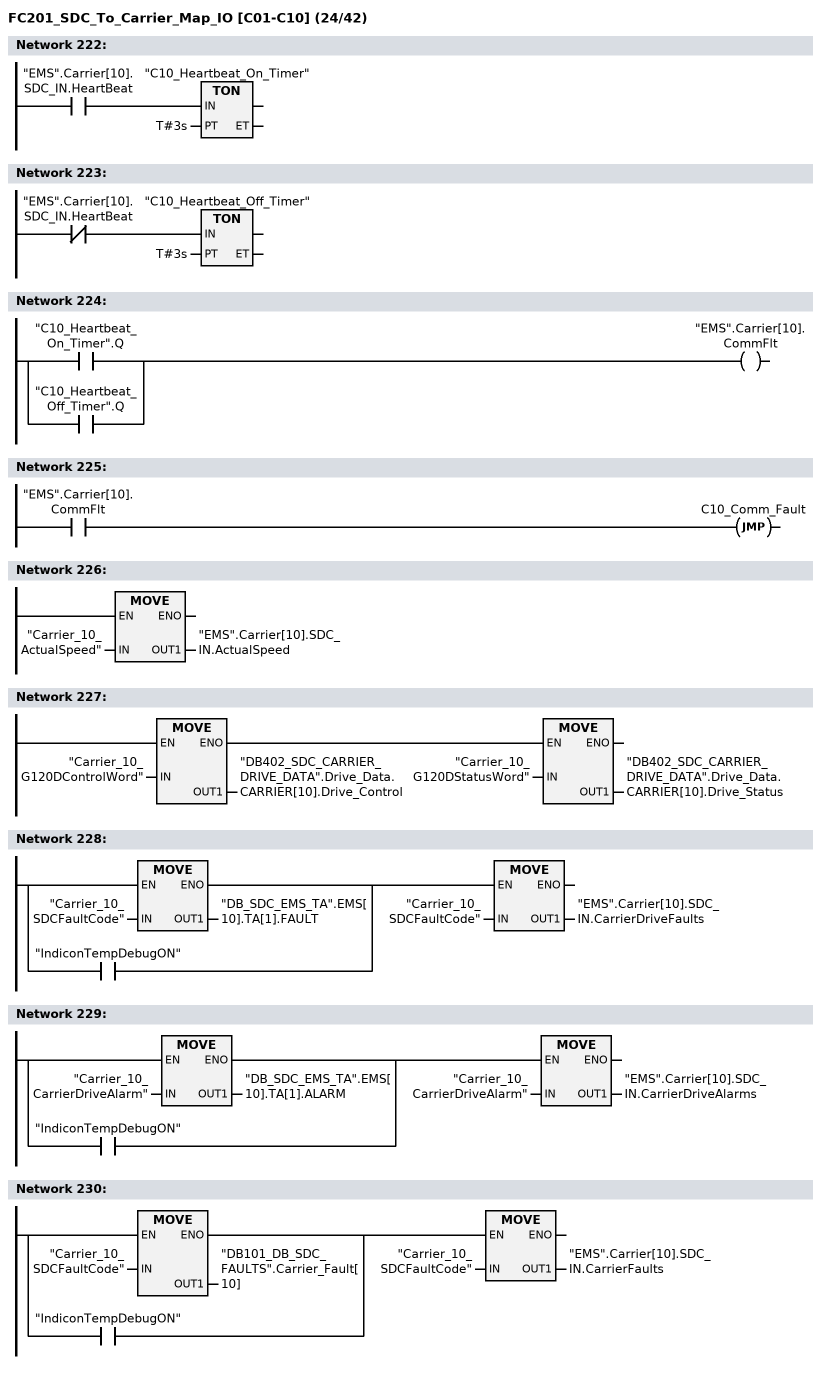
   "C10_Heartbeat_On_Timer".TON(IN := "EMS".Carrier[10].SDC_IN.HeartBeat, PT := T#3s);
END_REGION

REGION Network 223
   "C10_Heartbeat_Off_Timer".TON(IN := NOT "EMS".Carrier[10].SDC_IN.HeartBeat, PT := T#3s);
END_REGION

REGION Network 224
   RUNG wire#powerrail
      Contact( "C10_Heartbeat_On_Timer".Q )
      wire#w1
      Coil( "EMS".Carrier[10].CommFlt )
   END_RUNG
   RUNG wire#powerrail
      Contact( "C10_Heartbeat_Off_Timer".Q )
   END_RUNG wire#w1
   // the same network as SCL:
   "EMS".Carrier[10].CommFlt := "C10_Heartbeat_On_Timer".Q OR "C10_Heartbeat_Off_Timer".Q;
END_REGION

REGION Network 225
   RUNG wire#powerrail
      Contact( "EMS".Carrier[10].CommFlt )
      JumpCoil( C10_Comm_Fault )
   END_RUNG
   // the same network as SCL:
   IF "EMS".Carrier[10].CommFlt THEN GOTO C10_Comm_Fault; END_IF;
END_REGION

REGION Network 226
   RUNG wire#powerrail
      Move(in := "Carrier_10_ActualSpeed", out1 => "EMS".Carrier[10].SDC_IN.ActualSpeed)
   END_RUNG
   // the same network as SCL:
   "EMS".Carrier[10].SDC_IN.ActualSpeed := "Carrier_10_ActualSpeed";
END_REGION

REGION Network 227
   RUNG wire#powerrail
      Move(in := "Carrier_10_G120DControlWord", out1 => "DB402_SDC_CARRIER_DRIVE_DATA".Drive_Data.CARRIER[10].Drive_Control)
      Move(in := "Carrier_10_G120DStatusWord", out1 => "DB402_SDC_CARRIER_DRIVE_DATA".Drive_Data.CARRIER[10].Drive_Status)
   END_RUNG
   // the same network as SCL:
   "DB402_SDC_CARRIER_DRIVE_DATA".Drive_Data.CARRIER[10].Drive_Control := "Carrier_10_G120DControlWord";
   "DB402_SDC_CARRIER_DRIVE_DATA".Drive_Data.CARRIER[10].Drive_Status := "Carrier_10_G120DStatusWord";
END_REGION

REGION Network 228
   RUNG wire#powerrail
      Move(in := "Carrier_10_SDCFaultCode", out1 => "DB_SDC_EMS_TA".EMS[10].TA[1].FAULT)
      wire#w1
      Move(in := "Carrier_10_SDCFaultCode", out1 => "EMS".Carrier[10].SDC_IN.CarrierDriveFaults)
   END_RUNG
   RUNG wire#powerrail
      Contact( "IndiconTempDebugON" )
   END_RUNG wire#w1
   // the same network as SCL:
   "DB_SDC_EMS_TA".EMS[10].TA[1].FAULT := "Carrier_10_SDCFaultCode";
   IF TRUE OR "IndiconTempDebugON" THEN
       "EMS".Carrier[10].SDC_IN.CarrierDriveFaults := "Carrier_10_SDCFaultCode";
   END_IF;
END_REGION

REGION Network 229
   RUNG wire#powerrail
      Move(in := "Carrier_10_CarrierDriveAlarm", out1 => "DB_SDC_EMS_TA".EMS[10].TA[1].ALARM)
      wire#w1
      Move(in := "Carrier_10_CarrierDriveAlarm", out1 => "EMS".Carrier[10].SDC_IN.CarrierDriveAlarms)
   END_RUNG
   RUNG wire#powerrail
      Contact( "IndiconTempDebugON" )
   END_RUNG wire#w1
   // the same network as SCL:
   "DB_SDC_EMS_TA".EMS[10].TA[1].ALARM := "Carrier_10_CarrierDriveAlarm";
   IF TRUE OR "IndiconTempDebugON" THEN
       "EMS".Carrier[10].SDC_IN.CarrierDriveAlarms := "Carrier_10_CarrierDriveAlarm";
   END_IF;
END_REGION

REGION Network 230
   RUNG wire#powerrail
      Move(in := "Carrier_10_SDCFaultCode", out1 => "DB101_DB_SDC_FAULTS".Carrier_Fault[10])
      wire#w1
      Move(in := "Carrier_10_SDCFaultCode", out1 => "EMS".Carrier[10].SDC_IN.CarrierFaults)
   END_RUNG
   RUNG wire#powerrail
      Contact( "IndiconTempDebugON" )
   END_RUNG wire#w1
   // the same network as SCL:
   "DB101_DB_SDC_FAULTS".Carrier_Fault[10] := "Carrier_10_SDCFaultCode";
   IF TRUE OR "IndiconTempDebugON" THEN
       "EMS".Carrier[10].SDC_IN.CarrierFaults := "Carrier_10_SDCFaultCode";
   END_IF;
END_REGION

REGION Network 231
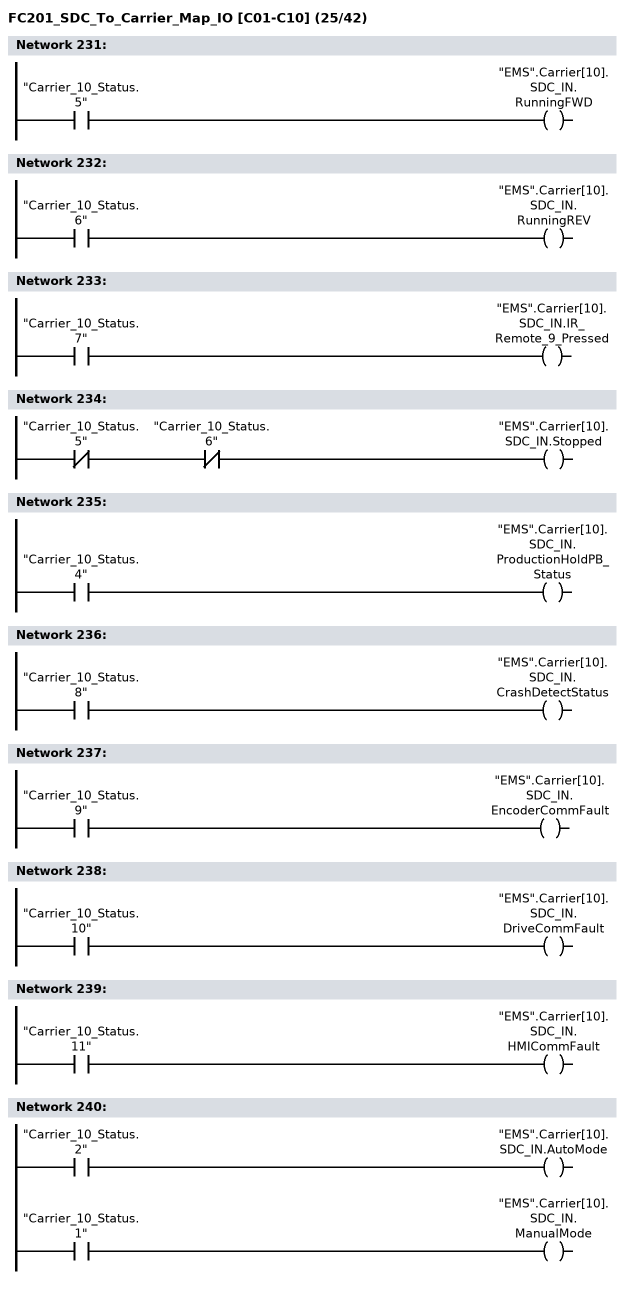
   RUNG wire#powerrail
      Contact( "Carrier_10_Status.5" )
      Coil( "EMS".Carrier[10].SDC_IN.RunningFWD )
   END_RUNG
   // the same network as SCL:
   "EMS".Carrier[10].SDC_IN.RunningFWD := "Carrier_10_Status.5";
END_REGION

REGION Network 232
   RUNG wire#powerrail
      Contact( "Carrier_10_Status.6" )
      Coil( "EMS".Carrier[10].SDC_IN.RunningREV )
   END_RUNG
   // the same network as SCL:
   "EMS".Carrier[10].SDC_IN.RunningREV := "Carrier_10_Status.6";
END_REGION

REGION Network 233
   RUNG wire#powerrail
      Contact( "Carrier_10_Status.7" )
      Coil( "EMS".Carrier[10].SDC_IN.IR_Remote_9_Pressed )
   END_RUNG
   // the same network as SCL:
   "EMS".Carrier[10].SDC_IN.IR_Remote_9_Pressed := "Carrier_10_Status.7";
END_REGION

REGION Network 234
   RUNG wire#powerrail
      I_Contact( "Carrier_10_Status.5" )
      I_Contact( "Carrier_10_Status.6" )
      Coil( "EMS".Carrier[10].SDC_IN.Stopped )
   END_RUNG
   // the same network as SCL:
   "EMS".Carrier[10].SDC_IN.Stopped := NOT "Carrier_10_Status.5" AND NOT "Carrier_10_Status.6";
END_REGION

REGION Network 235
   RUNG wire#powerrail
      Contact( "Carrier_10_Status.4" )
      Coil( "EMS".Carrier[10].SDC_IN.ProductionHoldPB_Status )
   END_RUNG
   // the same network as SCL:
   "EMS".Carrier[10].SDC_IN.ProductionHoldPB_Status := "Carrier_10_Status.4";
END_REGION

REGION Network 236
   RUNG wire#powerrail
      Contact( "Carrier_10_Status.8" )
      Coil( "EMS".Carrier[10].SDC_IN.CrashDetectStatus )
   END_RUNG
   // the same network as SCL:
   "EMS".Carrier[10].SDC_IN.CrashDetectStatus := "Carrier_10_Status.8";
END_REGION

REGION Network 237
   RUNG wire#powerrail
      Contact( "Carrier_10_Status.9" )
      Coil( "EMS".Carrier[10].SDC_IN.EncoderCommFault )
   END_RUNG
   // the same network as SCL:
   "EMS".Carrier[10].SDC_IN.EncoderCommFault := "Carrier_10_Status.9";
END_REGION

REGION Network 238
   RUNG wire#powerrail
      Contact( "Carrier_10_Status.10" )
      Coil( "EMS".Carrier[10].SDC_IN.DriveCommFault )
   END_RUNG
   // the same network as SCL:
   "EMS".Carrier[10].SDC_IN.DriveCommFault := "Carrier_10_Status.10";
END_REGION

REGION Network 239
   RUNG wire#powerrail
      Contact( "Carrier_10_Status.11" )
      Coil( "EMS".Carrier[10].SDC_IN.HMICommFault )
   END_RUNG
   // the same network as SCL:
   "EMS".Carrier[10].SDC_IN.HMICommFault := "Carrier_10_Status.11";
END_REGION

REGION Network 240
   RUNG wire#powerrail
      Contact( "Carrier_10_Status.2" )
      Coil( "EMS".Carrier[10].SDC_IN.AutoMode )
   END_RUNG
   RUNG wire#powerrail
      Contact( "Carrier_10_Status.1" )
      Coil( "EMS".Carrier[10].SDC_IN.ManualMode )
   END_RUNG
   // the same network as SCL:
   "EMS".Carrier[10].SDC_IN.AutoMode := "Carrier_10_Status.2";
   "EMS".Carrier[10].SDC_IN.ManualMode := "Carrier_10_Status.1";
END_REGION

REGION Network 241
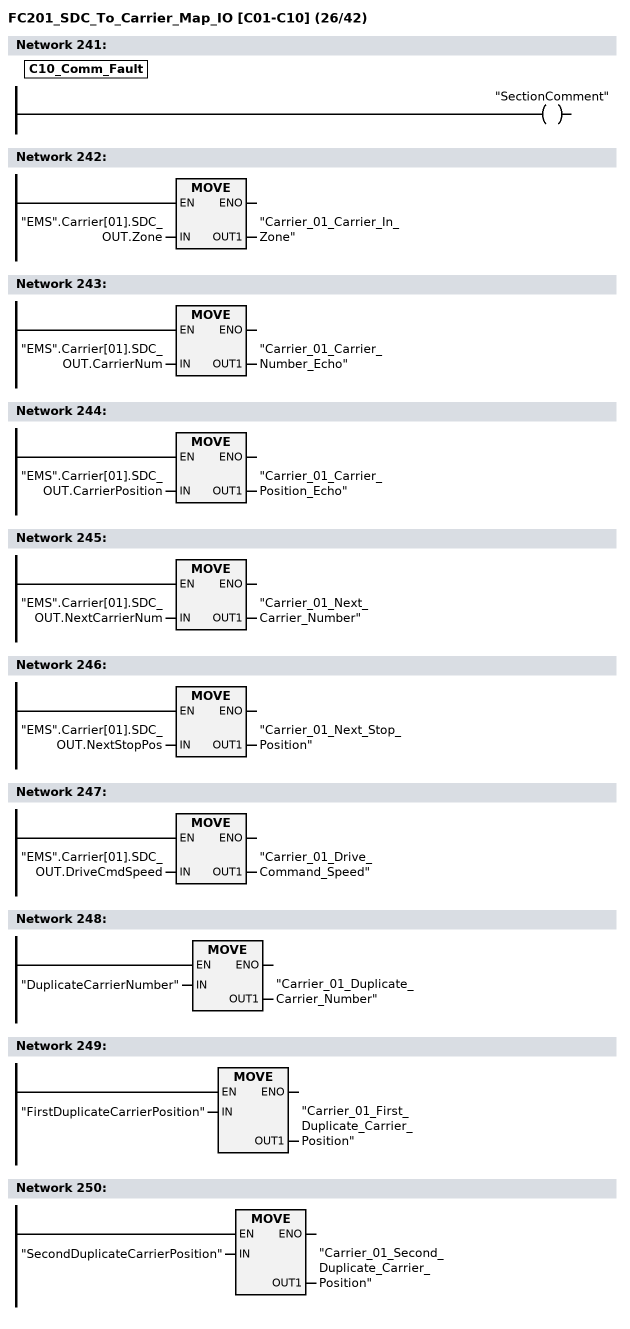
   Label( C10_Comm_Fault )
   RUNG wire#powerrail
      Coil( "SectionComment" )
   END_RUNG
   // the same network as SCL:
   C10_Comm_Fault:
   "SectionComment" := TRUE;
END_REGION

REGION Network 242
   RUNG wire#powerrail
      Move(in := "EMS".Carrier[01].SDC_OUT.Zone, out1 => "Carrier_01_Carrier_In_Zone")
   END_RUNG
   // the same network as SCL:
   "Carrier_01_Carrier_In_Zone" := "EMS".Carrier[01].SDC_OUT.Zone;
END_REGION

REGION Network 243
   RUNG wire#powerrail
      Move(in := "EMS".Carrier[01].SDC_OUT.CarrierNum, out1 => "Carrier_01_Carrier_Number_Echo")
   END_RUNG
   // the same network as SCL:
   "Carrier_01_Carrier_Number_Echo" := "EMS".Carrier[01].SDC_OUT.CarrierNum;
END_REGION

REGION Network 244
   RUNG wire#powerrail
      Move(in := "EMS".Carrier[01].SDC_OUT.CarrierPosition, out1 => "Carrier_01_Carrier_Position_Echo")
   END_RUNG
   // the same network as SCL:
   "Carrier_01_Carrier_Position_Echo" := "EMS".Carrier[01].SDC_OUT.CarrierPosition;
END_REGION

REGION Network 245
   RUNG wire#powerrail
      Move(in := "EMS".Carrier[01].SDC_OUT.NextCarrierNum, out1 => "Carrier_01_Next_Carrier_Number")
   END_RUNG
   // the same network as SCL:
   "Carrier_01_Next_Carrier_Number" := "EMS".Carrier[01].SDC_OUT.NextCarrierNum;
END_REGION

REGION Network 246
   RUNG wire#powerrail
      Move(in := "EMS".Carrier[01].SDC_OUT.NextStopPos, out1 => "Carrier_01_Next_Stop_Position")
   END_RUNG
   // the same network as SCL:
   "Carrier_01_Next_Stop_Position" := "EMS".Carrier[01].SDC_OUT.NextStopPos;
END_REGION

REGION Network 247
   RUNG wire#powerrail
      Move(in := "EMS".Carrier[01].SDC_OUT.DriveCmdSpeed, out1 => "Carrier_01_Drive_Command_Speed")
   END_RUNG
   // the same network as SCL:
   "Carrier_01_Drive_Command_Speed" := "EMS".Carrier[01].SDC_OUT.DriveCmdSpeed;
END_REGION

REGION Network 248
   RUNG wire#powerrail
      Move(in := "DuplicateCarrierNumber", out1 => "Carrier_01_Duplicate_Carrier_Number")
   END_RUNG
   // the same network as SCL:
   "Carrier_01_Duplicate_Carrier_Number" := "DuplicateCarrierNumber";
END_REGION

REGION Network 249
   RUNG wire#powerrail
      Move(in := "FirstDuplicateCarrierPosition", out1 => "Carrier_01_First_Duplicate_Carrier_Position")
   END_RUNG
   // the same network as SCL:
   "Carrier_01_First_Duplicate_Carrier_Position" := "FirstDuplicateCarrierPosition";
END_REGION

REGION Network 250
   RUNG wire#powerrail
      Move(in := "SecondDuplicateCarrierPosition", out1 => "Carrier_01_Second_Duplicate_Carrier_Position")
   END_RUNG
   // the same network as SCL:
   "Carrier_01_Second_Duplicate_Carrier_Position" := "SecondDuplicateCarrierPosition";
END_REGION

REGION Network 251
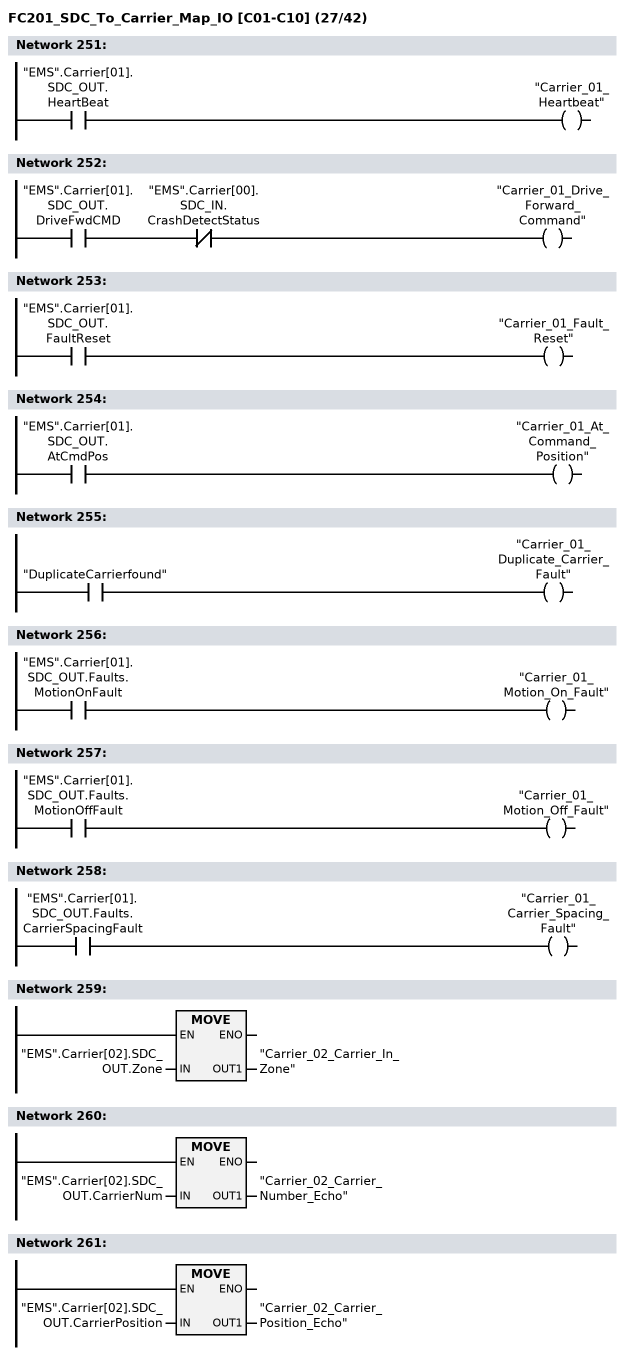
   RUNG wire#powerrail
      Contact( "EMS".Carrier[01].SDC_OUT.HeartBeat )
      Coil( "Carrier_01_Heartbeat" )
   END_RUNG
   // the same network as SCL:
   "Carrier_01_Heartbeat" := "EMS".Carrier[01].SDC_OUT.HeartBeat;
END_REGION

REGION Network 252
   RUNG wire#powerrail
      Contact( "EMS".Carrier[01].SDC_OUT.DriveFwdCMD )
      I_Contact( "EMS".Carrier[00].SDC_IN.CrashDetectStatus )
      Coil( "Carrier_01_Drive_Forward_Command" )
   END_RUNG
   // the same network as SCL:
   "Carrier_01_Drive_Forward_Command" := "EMS".Carrier[01].SDC_OUT.DriveFwdCMD AND NOT "EMS".Carrier[00].SDC_IN.CrashDetectStatus;
END_REGION

REGION Network 253
   RUNG wire#powerrail
      Contact( "EMS".Carrier[01].SDC_OUT.FaultReset )
      Coil( "Carrier_01_Fault_Reset" )
   END_RUNG
   // the same network as SCL:
   "Carrier_01_Fault_Reset" := "EMS".Carrier[01].SDC_OUT.FaultReset;
END_REGION

REGION Network 254
   RUNG wire#powerrail
      Contact( "EMS".Carrier[01].SDC_OUT.AtCmdPos )
      Coil( "Carrier_01_At_Command_Position" )
   END_RUNG
   // the same network as SCL:
   "Carrier_01_At_Command_Position" := "EMS".Carrier[01].SDC_OUT.AtCmdPos;
END_REGION

REGION Network 255
   RUNG wire#powerrail
      Contact( "DuplicateCarrierfound" )
      Coil( "Carrier_01_Duplicate_Carrier_Fault" )
   END_RUNG
   // the same network as SCL:
   "Carrier_01_Duplicate_Carrier_Fault" := "DuplicateCarrierfound";
END_REGION

REGION Network 256
   RUNG wire#powerrail
      Contact( "EMS".Carrier[01].SDC_OUT.Faults.MotionOnFault )
      Coil( "Carrier_01_Motion_On_Fault" )
   END_RUNG
   // the same network as SCL:
   "Carrier_01_Motion_On_Fault" := "EMS".Carrier[01].SDC_OUT.Faults.MotionOnFault;
END_REGION

REGION Network 257
   RUNG wire#powerrail
      Contact( "EMS".Carrier[01].SDC_OUT.Faults.MotionOffFault )
      Coil( "Carrier_01_Motion_Off_Fault" )
   END_RUNG
   // the same network as SCL:
   "Carrier_01_Motion_Off_Fault" := "EMS".Carrier[01].SDC_OUT.Faults.MotionOffFault;
END_REGION

REGION Network 258
   RUNG wire#powerrail
      Contact( "EMS".Carrier[01].SDC_OUT.Faults.CarrierSpacingFault )
      Coil( "Carrier_01_Carrier_Spacing_Fault" )
   END_RUNG
   // the same network as SCL:
   "Carrier_01_Carrier_Spacing_Fault" := "EMS".Carrier[01].SDC_OUT.Faults.CarrierSpacingFault;
END_REGION

REGION Network 259
   RUNG wire#powerrail
      Move(in := "EMS".Carrier[02].SDC_OUT.Zone, out1 => "Carrier_02_Carrier_In_Zone")
   END_RUNG
   // the same network as SCL:
   "Carrier_02_Carrier_In_Zone" := "EMS".Carrier[02].SDC_OUT.Zone;
END_REGION

REGION Network 260
   RUNG wire#powerrail
      Move(in := "EMS".Carrier[02].SDC_OUT.CarrierNum, out1 => "Carrier_02_Carrier_Number_Echo")
   END_RUNG
   // the same network as SCL:
   "Carrier_02_Carrier_Number_Echo" := "EMS".Carrier[02].SDC_OUT.CarrierNum;
END_REGION

REGION Network 261
   RUNG wire#powerrail
      Move(in := "EMS".Carrier[02].SDC_OUT.CarrierPosition, out1 => "Carrier_02_Carrier_Position_Echo")
   END_RUNG
   // the same network as SCL:
   "Carrier_02_Carrier_Position_Echo" := "EMS".Carrier[02].SDC_OUT.CarrierPosition;
END_REGION

REGION Network 262
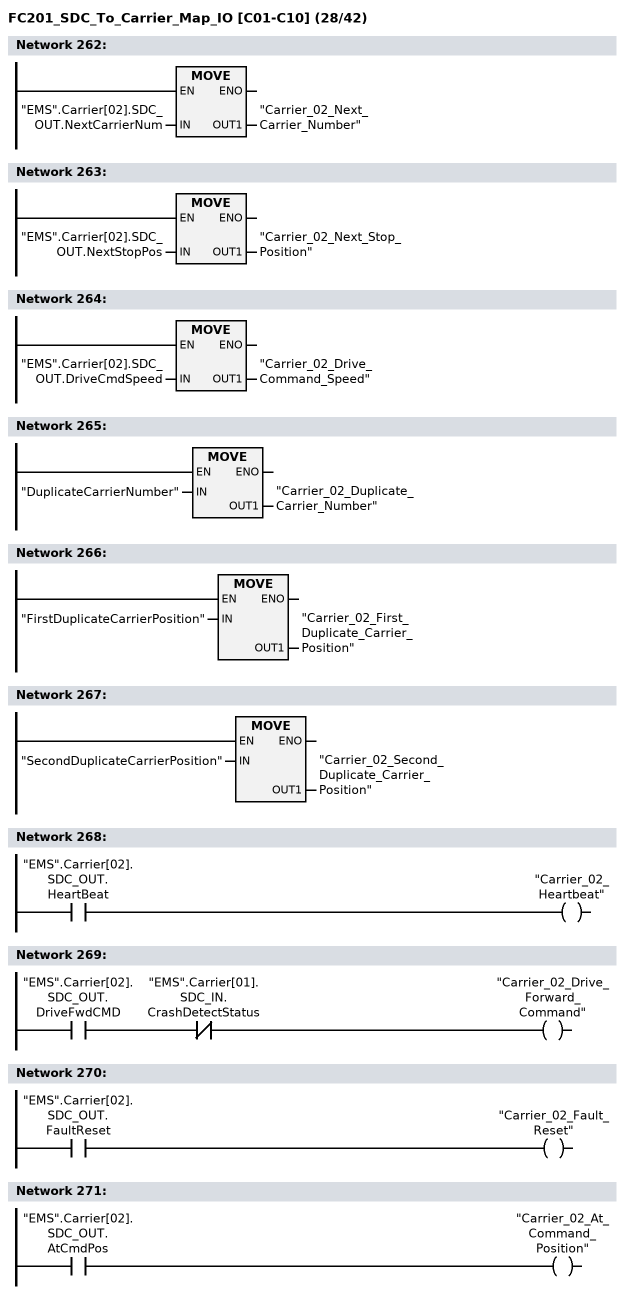
   RUNG wire#powerrail
      Move(in := "EMS".Carrier[02].SDC_OUT.NextCarrierNum, out1 => "Carrier_02_Next_Carrier_Number")
   END_RUNG
   // the same network as SCL:
   "Carrier_02_Next_Carrier_Number" := "EMS".Carrier[02].SDC_OUT.NextCarrierNum;
END_REGION

REGION Network 263
   RUNG wire#powerrail
      Move(in := "EMS".Carrier[02].SDC_OUT.NextStopPos, out1 => "Carrier_02_Next_Stop_Position")
   END_RUNG
   // the same network as SCL:
   "Carrier_02_Next_Stop_Position" := "EMS".Carrier[02].SDC_OUT.NextStopPos;
END_REGION

REGION Network 264
   RUNG wire#powerrail
      Move(in := "EMS".Carrier[02].SDC_OUT.DriveCmdSpeed, out1 => "Carrier_02_Drive_Command_Speed")
   END_RUNG
   // the same network as SCL:
   "Carrier_02_Drive_Command_Speed" := "EMS".Carrier[02].SDC_OUT.DriveCmdSpeed;
END_REGION

REGION Network 265
   RUNG wire#powerrail
      Move(in := "DuplicateCarrierNumber", out1 => "Carrier_02_Duplicate_Carrier_Number")
   END_RUNG
   // the same network as SCL:
   "Carrier_02_Duplicate_Carrier_Number" := "DuplicateCarrierNumber";
END_REGION

REGION Network 266
   RUNG wire#powerrail
      Move(in := "FirstDuplicateCarrierPosition", out1 => "Carrier_02_First_Duplicate_Carrier_Position")
   END_RUNG
   // the same network as SCL:
   "Carrier_02_First_Duplicate_Carrier_Position" := "FirstDuplicateCarrierPosition";
END_REGION

REGION Network 267
   RUNG wire#powerrail
      Move(in := "SecondDuplicateCarrierPosition", out1 => "Carrier_02_Second_Duplicate_Carrier_Position")
   END_RUNG
   // the same network as SCL:
   "Carrier_02_Second_Duplicate_Carrier_Position" := "SecondDuplicateCarrierPosition";
END_REGION

REGION Network 268
   RUNG wire#powerrail
      Contact( "EMS".Carrier[02].SDC_OUT.HeartBeat )
      Coil( "Carrier_02_Heartbeat" )
   END_RUNG
   // the same network as SCL:
   "Carrier_02_Heartbeat" := "EMS".Carrier[02].SDC_OUT.HeartBeat;
END_REGION

REGION Network 269
   RUNG wire#powerrail
      Contact( "EMS".Carrier[02].SDC_OUT.DriveFwdCMD )
      I_Contact( "EMS".Carrier[01].SDC_IN.CrashDetectStatus )
      Coil( "Carrier_02_Drive_Forward_Command" )
   END_RUNG
   // the same network as SCL:
   "Carrier_02_Drive_Forward_Command" := "EMS".Carrier[02].SDC_OUT.DriveFwdCMD AND NOT "EMS".Carrier[01].SDC_IN.CrashDetectStatus;
END_REGION

REGION Network 270
   RUNG wire#powerrail
      Contact( "EMS".Carrier[02].SDC_OUT.FaultReset )
      Coil( "Carrier_02_Fault_Reset" )
   END_RUNG
   // the same network as SCL:
   "Carrier_02_Fault_Reset" := "EMS".Carrier[02].SDC_OUT.FaultReset;
END_REGION

REGION Network 271
   RUNG wire#powerrail
      Contact( "EMS".Carrier[02].SDC_OUT.AtCmdPos )
      Coil( "Carrier_02_At_Command_Position" )
   END_RUNG
   // the same network as SCL:
   "Carrier_02_At_Command_Position" := "EMS".Carrier[02].SDC_OUT.AtCmdPos;
END_REGION

REGION Network 272
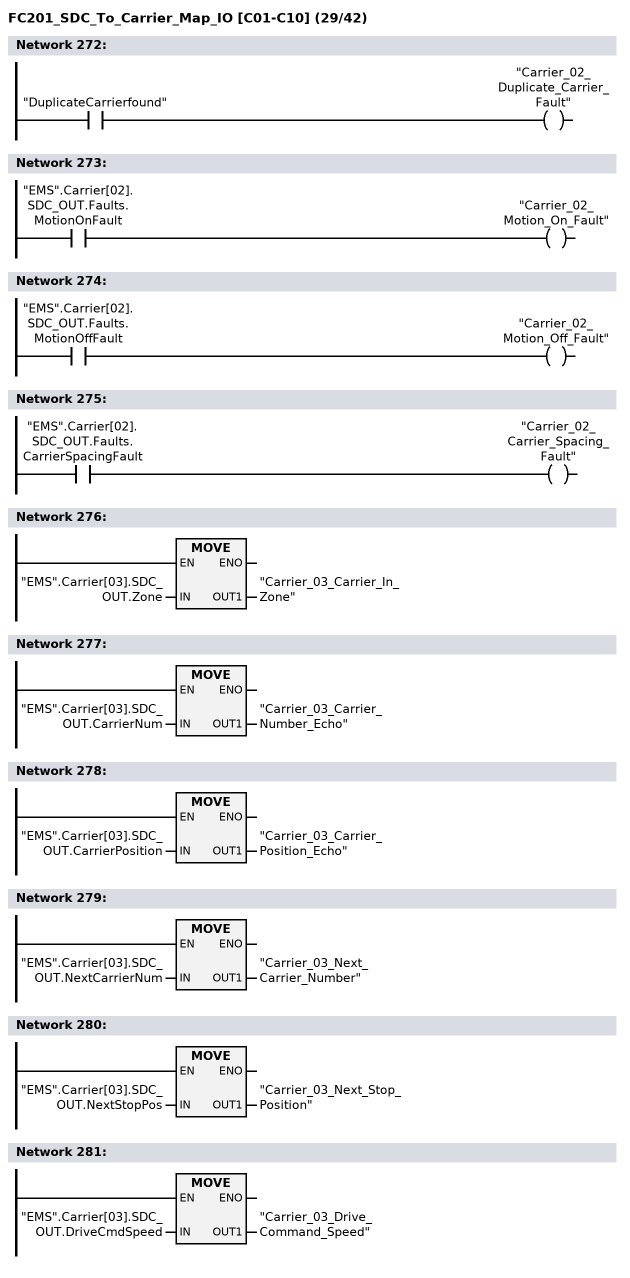
   RUNG wire#powerrail
      Contact( "DuplicateCarrierfound" )
      Coil( "Carrier_02_Duplicate_Carrier_Fault" )
   END_RUNG
   // the same network as SCL:
   "Carrier_02_Duplicate_Carrier_Fault" := "DuplicateCarrierfound";
END_REGION

REGION Network 273
   RUNG wire#powerrail
      Contact( "EMS".Carrier[02].SDC_OUT.Faults.MotionOnFault )
      Coil( "Carrier_02_Motion_On_Fault" )
   END_RUNG
   // the same network as SCL:
   "Carrier_02_Motion_On_Fault" := "EMS".Carrier[02].SDC_OUT.Faults.MotionOnFault;
END_REGION

REGION Network 274
   RUNG wire#powerrail
      Contact( "EMS".Carrier[02].SDC_OUT.Faults.MotionOffFault )
      Coil( "Carrier_02_Motion_Off_Fault" )
   END_RUNG
   // the same network as SCL:
   "Carrier_02_Motion_Off_Fault" := "EMS".Carrier[02].SDC_OUT.Faults.MotionOffFault;
END_REGION

REGION Network 275
   RUNG wire#powerrail
      Contact( "EMS".Carrier[02].SDC_OUT.Faults.CarrierSpacingFault )
      Coil( "Carrier_02_Carrier_Spacing_Fault" )
   END_RUNG
   // the same network as SCL:
   "Carrier_02_Carrier_Spacing_Fault" := "EMS".Carrier[02].SDC_OUT.Faults.CarrierSpacingFault;
END_REGION

REGION Network 276
   RUNG wire#powerrail
      Move(in := "EMS".Carrier[03].SDC_OUT.Zone, out1 => "Carrier_03_Carrier_In_Zone")
   END_RUNG
   // the same network as SCL:
   "Carrier_03_Carrier_In_Zone" := "EMS".Carrier[03].SDC_OUT.Zone;
END_REGION

REGION Network 277
   RUNG wire#powerrail
      Move(in := "EMS".Carrier[03].SDC_OUT.CarrierNum, out1 => "Carrier_03_Carrier_Number_Echo")
   END_RUNG
   // the same network as SCL:
   "Carrier_03_Carrier_Number_Echo" := "EMS".Carrier[03].SDC_OUT.CarrierNum;
END_REGION

REGION Network 278
   RUNG wire#powerrail
      Move(in := "EMS".Carrier[03].SDC_OUT.CarrierPosition, out1 => "Carrier_03_Carrier_Position_Echo")
   END_RUNG
   // the same network as SCL:
   "Carrier_03_Carrier_Position_Echo" := "EMS".Carrier[03].SDC_OUT.CarrierPosition;
END_REGION

REGION Network 279
   RUNG wire#powerrail
      Move(in := "EMS".Carrier[03].SDC_OUT.NextCarrierNum, out1 => "Carrier_03_Next_Carrier_Number")
   END_RUNG
   // the same network as SCL:
   "Carrier_03_Next_Carrier_Number" := "EMS".Carrier[03].SDC_OUT.NextCarrierNum;
END_REGION

REGION Network 280
   RUNG wire#powerrail
      Move(in := "EMS".Carrier[03].SDC_OUT.NextStopPos, out1 => "Carrier_03_Next_Stop_Position")
   END_RUNG
   // the same network as SCL:
   "Carrier_03_Next_Stop_Position" := "EMS".Carrier[03].SDC_OUT.NextStopPos;
END_REGION

REGION Network 281
   RUNG wire#powerrail
      Move(in := "EMS".Carrier[03].SDC_OUT.DriveCmdSpeed, out1 => "Carrier_03_Drive_Command_Speed")
   END_RUNG
   // the same network as SCL:
   "Carrier_03_Drive_Command_Speed" := "EMS".Carrier[03].SDC_OUT.DriveCmdSpeed;
END_REGION

REGION Network 282
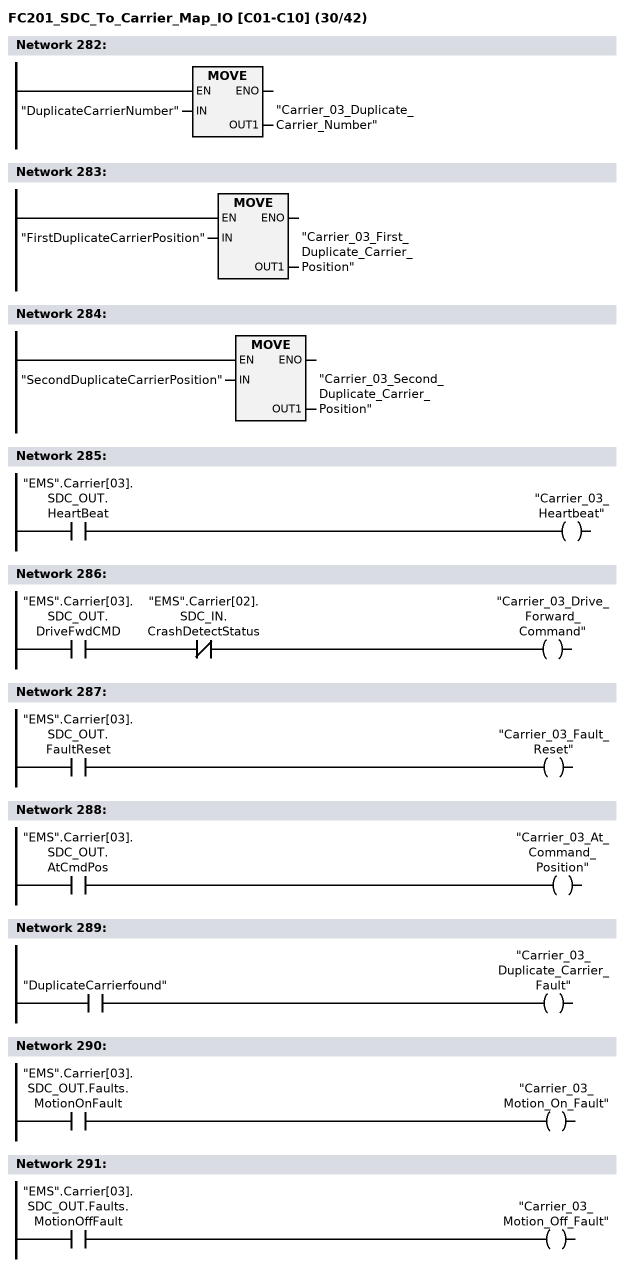
   RUNG wire#powerrail
      Move(in := "DuplicateCarrierNumber", out1 => "Carrier_03_Duplicate_Carrier_Number")
   END_RUNG
   // the same network as SCL:
   "Carrier_03_Duplicate_Carrier_Number" := "DuplicateCarrierNumber";
END_REGION

REGION Network 283
   RUNG wire#powerrail
      Move(in := "FirstDuplicateCarrierPosition", out1 => "Carrier_03_First_Duplicate_Carrier_Position")
   END_RUNG
   // the same network as SCL:
   "Carrier_03_First_Duplicate_Carrier_Position" := "FirstDuplicateCarrierPosition";
END_REGION

REGION Network 284
   RUNG wire#powerrail
      Move(in := "SecondDuplicateCarrierPosition", out1 => "Carrier_03_Second_Duplicate_Carrier_Position")
   END_RUNG
   // the same network as SCL:
   "Carrier_03_Second_Duplicate_Carrier_Position" := "SecondDuplicateCarrierPosition";
END_REGION

REGION Network 285
   RUNG wire#powerrail
      Contact( "EMS".Carrier[03].SDC_OUT.HeartBeat )
      Coil( "Carrier_03_Heartbeat" )
   END_RUNG
   // the same network as SCL:
   "Carrier_03_Heartbeat" := "EMS".Carrier[03].SDC_OUT.HeartBeat;
END_REGION

REGION Network 286
   RUNG wire#powerrail
      Contact( "EMS".Carrier[03].SDC_OUT.DriveFwdCMD )
      I_Contact( "EMS".Carrier[02].SDC_IN.CrashDetectStatus )
      Coil( "Carrier_03_Drive_Forward_Command" )
   END_RUNG
   // the same network as SCL:
   "Carrier_03_Drive_Forward_Command" := "EMS".Carrier[03].SDC_OUT.DriveFwdCMD AND NOT "EMS".Carrier[02].SDC_IN.CrashDetectStatus;
END_REGION

REGION Network 287
   RUNG wire#powerrail
      Contact( "EMS".Carrier[03].SDC_OUT.FaultReset )
      Coil( "Carrier_03_Fault_Reset" )
   END_RUNG
   // the same network as SCL:
   "Carrier_03_Fault_Reset" := "EMS".Carrier[03].SDC_OUT.FaultReset;
END_REGION

REGION Network 288
   RUNG wire#powerrail
      Contact( "EMS".Carrier[03].SDC_OUT.AtCmdPos )
      Coil( "Carrier_03_At_Command_Position" )
   END_RUNG
   // the same network as SCL:
   "Carrier_03_At_Command_Position" := "EMS".Carrier[03].SDC_OUT.AtCmdPos;
END_REGION

REGION Network 289
   RUNG wire#powerrail
      Contact( "DuplicateCarrierfound" )
      Coil( "Carrier_03_Duplicate_Carrier_Fault" )
   END_RUNG
   // the same network as SCL:
   "Carrier_03_Duplicate_Carrier_Fault" := "DuplicateCarrierfound";
END_REGION

REGION Network 290
   RUNG wire#powerrail
      Contact( "EMS".Carrier[03].SDC_OUT.Faults.MotionOnFault )
      Coil( "Carrier_03_Motion_On_Fault" )
   END_RUNG
   // the same network as SCL:
   "Carrier_03_Motion_On_Fault" := "EMS".Carrier[03].SDC_OUT.Faults.MotionOnFault;
END_REGION

REGION Network 291
   RUNG wire#powerrail
      Contact( "EMS".Carrier[03].SDC_OUT.Faults.MotionOffFault )
      Coil( "Carrier_03_Motion_Off_Fault" )
   END_RUNG
   // the same network as SCL:
   "Carrier_03_Motion_Off_Fault" := "EMS".Carrier[03].SDC_OUT.Faults.MotionOffFault;
END_REGION

REGION Network 292
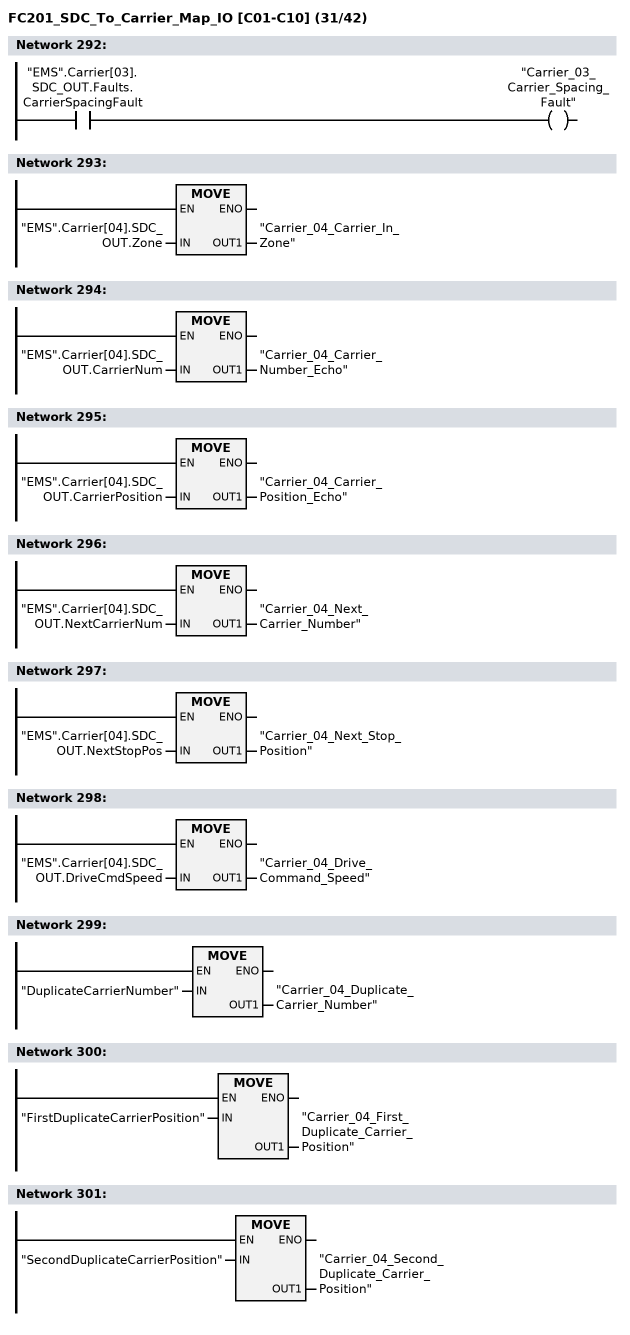
   RUNG wire#powerrail
      Contact( "EMS".Carrier[03].SDC_OUT.Faults.CarrierSpacingFault )
      Coil( "Carrier_03_Carrier_Spacing_Fault" )
   END_RUNG
   // the same network as SCL:
   "Carrier_03_Carrier_Spacing_Fault" := "EMS".Carrier[03].SDC_OUT.Faults.CarrierSpacingFault;
END_REGION

REGION Network 293
   RUNG wire#powerrail
      Move(in := "EMS".Carrier[04].SDC_OUT.Zone, out1 => "Carrier_04_Carrier_In_Zone")
   END_RUNG
   // the same network as SCL:
   "Carrier_04_Carrier_In_Zone" := "EMS".Carrier[04].SDC_OUT.Zone;
END_REGION

REGION Network 294
   RUNG wire#powerrail
      Move(in := "EMS".Carrier[04].SDC_OUT.CarrierNum, out1 => "Carrier_04_Carrier_Number_Echo")
   END_RUNG
   // the same network as SCL:
   "Carrier_04_Carrier_Number_Echo" := "EMS".Carrier[04].SDC_OUT.CarrierNum;
END_REGION

REGION Network 295
   RUNG wire#powerrail
      Move(in := "EMS".Carrier[04].SDC_OUT.CarrierPosition, out1 => "Carrier_04_Carrier_Position_Echo")
   END_RUNG
   // the same network as SCL:
   "Carrier_04_Carrier_Position_Echo" := "EMS".Carrier[04].SDC_OUT.CarrierPosition;
END_REGION

REGION Network 296
   RUNG wire#powerrail
      Move(in := "EMS".Carrier[04].SDC_OUT.NextCarrierNum, out1 => "Carrier_04_Next_Carrier_Number")
   END_RUNG
   // the same network as SCL:
   "Carrier_04_Next_Carrier_Number" := "EMS".Carrier[04].SDC_OUT.NextCarrierNum;
END_REGION

REGION Network 297
   RUNG wire#powerrail
      Move(in := "EMS".Carrier[04].SDC_OUT.NextStopPos, out1 => "Carrier_04_Next_Stop_Position")
   END_RUNG
   // the same network as SCL:
   "Carrier_04_Next_Stop_Position" := "EMS".Carrier[04].SDC_OUT.NextStopPos;
END_REGION

REGION Network 298
   RUNG wire#powerrail
      Move(in := "EMS".Carrier[04].SDC_OUT.DriveCmdSpeed, out1 => "Carrier_04_Drive_Command_Speed")
   END_RUNG
   // the same network as SCL:
   "Carrier_04_Drive_Command_Speed" := "EMS".Carrier[04].SDC_OUT.DriveCmdSpeed;
END_REGION

REGION Network 299
   RUNG wire#powerrail
      Move(in := "DuplicateCarrierNumber", out1 => "Carrier_04_Duplicate_Carrier_Number")
   END_RUNG
   // the same network as SCL:
   "Carrier_04_Duplicate_Carrier_Number" := "DuplicateCarrierNumber";
END_REGION

REGION Network 300
   RUNG wire#powerrail
      Move(in := "FirstDuplicateCarrierPosition", out1 => "Carrier_04_First_Duplicate_Carrier_Position")
   END_RUNG
   // the same network as SCL:
   "Carrier_04_First_Duplicate_Carrier_Position" := "FirstDuplicateCarrierPosition";
END_REGION

REGION Network 301
   RUNG wire#powerrail
      Move(in := "SecondDuplicateCarrierPosition", out1 => "Carrier_04_Second_Duplicate_Carrier_Position")
   END_RUNG
   // the same network as SCL:
   "Carrier_04_Second_Duplicate_Carrier_Position" := "SecondDuplicateCarrierPosition";
END_REGION

REGION Network 302